// TIA Portal project "Delta_Praktika_P&P" (V17)

(* hardware
DEVICE "S7-1500/ET200MP station_1"  S7-1500 station
   slot 0: "Rail_0"  Rack  6ES7 590-1***0-0AA0
   slot 1: "PLC_2"  CPU 1517TF-3 PN/DP  6ES7 517-3UP00-0AB0  V2.9
      slot 3: "CPU display_1"  6ES7591-1BA00-0AA0
      slot 32768: "PROFINET interface_1"  X1
      slot 33024: "PROFINET interface_2"  X2
      slot 33280: "DP interface_1"  X3
      slot 34817: "Virtual CP interface port_1"  Virtual CP interface port  Virtual CP interface port
DEVICE "ET 200SP station_1"  ET 200SP-Station
   slot 0: "Rack_0"  Rack  6ES5 710-8MAx1
   slot 0: "et200sp"  IM 155-6 PN/2 HF  6ES7 155-6AU01-0CN0  V4.2
   slot 1: "DI 8x24VDC HF_1"  DI 8x24VDC HF  6ES7 131-6BF00-0CA0  V2.0
      slot 1: "DI 8x24VDC HF_1"  DI 8x24VDC HF
   slot 2: "DQ 8x24VDC/0.5A HF_1"  DQ 8x24VDC/0.5A HF  6ES7 132-6BF00-0CA0  V2.0
      slot 1: "DQ 8x24VDC/0.5A HF_1"  DQ 8x24VDC/0.5A HF
   slot 3: "CM 4xIO-Link_1"  CM 4xIO-Link  6ES7 137-6BD00-0BA0  V2.2
      slot 1: "CM 4xIO-Link_1"  6ES7 137-6BD00-0BA0
   slot 4: "Server module_1"  Server module  6ES7 193-6PA00-0AA0  V1.1
      slot 1: "Server module_1"  Server module
   slot 127: "BA 2xRJ45"  BA 2xRJ45  6ES7 193-6AR00-0AA0  V0.0
      slot 1: "Port_1"  X1 P1 R  6ES7 193-6AR00-0AA0  V0.0
      slot 2: "Port_2"  X1 P2 R  6ES7 193-6AR00-0AA0  V0.0
DEVICE "SINAMICS V_1"  SINAMICS V
   slot 0: "SINAMICS V90 PN Rack"  Rail  1.0
   slot 0: "a1"  V90 PN  6SL3 210-5FB10-4UFx  V1.4
      slot 1: "Drive object"  Drive Object
         slot 1: "Module access point"  Module Access Point
         slot 2: "Without PROFIsafe"  No ProfiSafe
         slot 3: "Telegram"  SIEMENS Telegramm 105
DEVICE "SINAMICS V_2"  SINAMICS V
   slot 0: "SINAMICS V90 PN Rack"  Rail  1.0
   slot 0: "a3"  V90 PN  6SL3 210-5FB10-4UFx  V1.4
      slot 1: "Drive object"  Drive Object
         slot 1: "Module access point"  Module Access Point
         slot 2: "Without PROFIsafe"  No ProfiSafe
         slot 3: "Telegram"  SIEMENS Telegramm 105
DEVICE "SINAMICS V_3"  SINAMICS V
   slot 0: "SINAMICS V90 PN Rack"  Rail  1.0
   slot 0: "a2"  V90 PN  6SL3 210-5FB10-4UFx  V1.4
      slot 1: "Drive object"  Drive Object
         slot 1: "Module access point"  Module Access Point
         slot 2: "Without PROFIsafe"  No ProfiSafe
         slot 3: "Telegram"  SIEMENS Telegramm 105
DEVICE "HMI_1"  KTP1200 Basic PN
   slot 0: "HMI_1"  KTP1200 Basic PN  6AV2 123-2MB03-0AX0  17.0.0.0
   slot 1: "HMI_RT_1"  KTP1200 Basic PN  6AV2 123-2MB03-0AX0  17.0.0.0
   slot 5: "HMI_1.IE_CP_1"  PROFINET Interface  17.0.0.0
      slot 1: "Interfaz PROFINET_1"  PROFINET Interface
         slot 1: "Port_1"  Port
*)

// ===== PLC "PLC_2"  CPU 1517TF-3 PN/DP =====

VAR_GLOBAL   // PLC tag table "Default tag table"
   "A1_Actor_Interface_AddressIn" AT %I0.0 : "PD_TEL3_IN";
   "A1_Actor_Interface_AddressOut" AT %Q0.0 : "PD_TEL3_OUT";
   "A2_Actor_Interface_AddressIn" AT %I18.0 : "PD_TEL3_IN";
   "A2_Actor_Interface_AddressOut" AT %Q10.0 : "PD_TEL3_OUT";
   "A3_Actor_Interface_AddressIn" AT %I36.0 : "PD_TEL3_IN";
   "A3_Actor_Interface_AddressOut" AT %Q20.0 : "PD_TEL3_OUT";
   "A1_axis_Actor_Interface_AddressIn" AT %I0.0 : "PD_TEL105_IN";
   "A1_axis_Actor_Interface_AddressOut" AT %Q0.0 : "PD_TEL105_OUT";
   "a2_axis_Actor_Interface_AddressIn" AT %I20.0 : "PD_TEL105_IN";
   "a2_axis_Actor_Interface_AddressOut" AT %Q63.0 : "PD_TEL105_OUT";
   "a3_asix_Actor_Interface_AddressIn" AT %I87.0 : "PD_TEL105_IN";
   "a3_asix_Actor_Interface_AddressOut" AT %Q83.0 : "PD_TEL105_OUT";
   "Freno_a1" AT %Q30.1 : Bool;
   "marka_Freno_a1" AT %M30.1 : Bool;
   "marka_Freno_a2" AT %M30.2 : Bool;
   "Freno_a2" AT %Q30.2 : Bool;
   "Freno_a3" AT %Q30.0 : Bool;
   "marka_Freno_a3" AT %M30.0 : Bool;
   "System_Byte" AT %MB256 : Byte;
   "FirstScan" AT %M256.0 : Bool;
   "DiagStatusUpdate" AT %M256.1 : Bool;
   "AlwaysTRUE" AT %M256.2 : Bool;
   "AlwaysFALSE" AT %M256.3 : Bool;
   "Clock_Byte" AT %MB255 : Byte;
   "Clock_10Hz" AT %M255.0 : Bool;
   "Clock_5Hz" AT %M255.1 : Bool;
   "Clock_2.5Hz" AT %M255.2 : Bool;
   "Clock_2Hz" AT %M255.3 : Bool;
   "Clock_1.25Hz" AT %M255.4 : Bool;
   "Clock_1Hz" AT %M255.5 : Bool;
   "Clock_0.625Hz" AT %M255.6 : Bool;
   "Clock_0.5Hz" AT %M255.7 : Bool;
   "Tag_1" AT %M401.0 : Bool;
   "JogFordward" AT %M150.0 : Bool;
   "JogBackward" AT %M150.1 : Bool;
   "Direction" AT %MB151 : USInt;
   "x+" AT %M152.0 : Bool;
   "x-" AT %M152.1 : Bool;
   "y+" AT %M152.2 : Bool;
   "y-" AT %M152.3 : Bool;
   "z+" AT %M152.4 : Bool;
   "z-" AT %M152.5 : Bool;
   "HABILITAR" AT %M150.2 : Bool;
   "Etapa0" AT %M0.0 : Bool;
   "HMI_start" AT %M10.0 : Bool;
   "Etapa1" AT %M0.1 : Bool;
   "Etapa2" AT %M0.2 : Bool;
   "Etapa3" AT %M0.3 : Bool;
   "Etapa4" AT %M0.4 : Bool;
   "Etapa5" AT %M0.5 : Bool;
   "Etapa6" AT %M0.6 : Bool;
   "Etapa7" AT %M0.7 : Bool;
   "kontagailua" AT %MW2 : Int;
   "Tag_2" AT %MB0 : Byte;
   "Tag_3" AT %M11.0 : Bool;
   "Etapa8" AT %M1.0 : Bool;
   "Etapa9" AT %M1.1 : Bool;
   "Etapa10" AT %M1.2 : Bool;
   "Etapa11" AT %M1.3 : Bool;
   "Etapa12" AT %M1.4 : Bool;
   "Tag_4" AT %MB1 : Byte;
   "Bentosa" AT %Q30.3 : Bool;
   "Tag_5" AT %M11.1 : Bool;
   "Tag_6" AT %M11.2 : Bool;
   "Tag_7" AT %M11.3 : Bool;
   "Tag_8" AT %M11.4 : Bool;
   "Tag_9" AT %M11.5 : Bool;
   "Tag_10" AT %M11.6 : Bool;
   "Tag_11" AT %M11.7 : Bool;
   "Tag_12" AT %M12.0 : Bool;
   "Tag_13" AT %M17.0 : Bool;
   "Tag_14" AT %M17.1 : Bool;
   "Tag_15" AT %M17.3 : Bool;
   "Tag_16" AT %M17.4 : Bool;
   "Tag_17" AT %M17.5 : Bool;
   "Tag_18" AT %M17.6 : Bool;
   "Tag_19" AT %M18.0 : Bool;
   "Tag_20" AT %M18.1 : Bool;
   "Tag_21" AT %M18.2 : Bool;
   "Tag_22" AT %M18.3 : Bool;
   "Tag_23" AT %M18.4 : Bool;
   "Tag_24" AT %M18.5 : Bool;
END_VAR

TYPE "LKinCtrl_typePathDynamics"
   STRUCT
      velocity : LReal := -1.0;   // >0.0: configured value used; <0.0: default TO setting used; for cmdType = 100 ==> waitTime in ms
      acceleration : LReal := -1.0;   // >0.0: configured value used; <0.0: default TO setting used
      deceleration : LReal := -1.0;   // >0.0: configured value used; <0.0: default TO setting used
      jerk : LReal := -1.0;   // >0.0: configured value used; <0.0: default TO setting used
   END_STRUCT;
END_TYPE

TYPE "LKinCtrl_typeSPTPDynamics"
   STRUCT
      velocityFactor : LReal;   // Factor for the velocity of axis movements in relation to the respective maximum velocity of the axes. Permitted value range: -1.0 < Factor ≤ 1.0
      accelerationFactor : LReal;   // Factor for the acceleration of axis movements in relation to the respective maximum acceleration of the axis. Permitted value range: -1.0 < Factor ≤ 1.0
      decelerationFactor : LReal;   // Factor for the deceleration of the axis movements in relation to the respective maximum deceleration of the axis. Permitted value range: -1.0 < Factor ≤ 1.0
      jerkFactor : LReal;   // Factor for the jerk of axis movements in relation to the respective maximum jerk of the axis. Permitted value range: -1.0 <Factor ≤ 0.0 and 0.1 < Factor ≤ 0.9
   END_STRUCT;
END_TYPE

TYPE "LKinCtrl_typeJogFrameDiagnostics"
VERSION : 0.1
// support: tech.team.motioncontrol@siemens.com
   STRUCT
      timeStamp : Date_And_Time;   // Time stamp at which the error occurred
      status : Word;   // Status of FB when error occurred
      stateNumber : DInt;   // State in the state machine of the FB when the error occurred
   END_STRUCT;
END_TYPE

TYPE "LKinCtrl_typeCartesianPosition"
   STRUCT
      x : LReal;   // X
      y : LReal;   // Y
      z : LReal;   // Z
      "a" : LReal;   // A
      "b" : LReal;   // B
      c : LReal;   // C
   END_STRUCT;
END_TYPE

TYPE "LKinCtrl_typeDynamics"
VERSION : 0.1
   STRUCT
      path : "LKinCtrl_typePathDynamics";   // Specification of the path dynamics
      orientation : "LKinCtrl_typePathDynamics";   // Specification of the orientation dynamics
      dynamicAdaption : DInt := 1;   // 0=no dynamic adaption, 1=dynamic adaptation with segmentation of the path, 2=dynamic adaptation without segmentation of the path
      directionA : DInt := 3;   // 1=positive direction, 2=negative direction, 3=shortest distance
      sPTP : "LKinCtrl_typeSPTPDynamics";   // Specification of the dynamic factor for sptp movement
   END_STRUCT;
END_TYPE

DATA_BLOCK "Power_DB"   // DB9
{ S7_Optimized_Access := 'TRUE' }
VERSION : 0.1
// stored: InstanceOfName Power
"Power"
BEGIN
END_DATA_BLOCK

DATA_BLOCK "Parametroak"   // DB11
{ S7_Optimized_Access := 'TRUE' }
VERSION : 0.1
   VAR
      Abiadura : LReal := 2.0;
      Azelerazioa : LReal := 40.0;
      Desazelerazioa : LReal := 40.0;
      Jerk : LReal := 400.0;
      offset : LReal := 30.0;
   END_VAR
BEGIN
END_DATA_BLOCK

DATA_BLOCK "Jog_DB"   // DB14
{ S7_Optimized_Access := 'TRUE' }
VERSION : 0.1
// stored: InstanceOfName Jog
"Jog"
BEGIN
END_DATA_BLOCK

DATA_BLOCK "Hominga_DB"   // DB18
{ S7_Optimized_Access := 'TRUE' }
VERSION : 0.1
// stored: InstanceOfName Hominga
"Hominga"
BEGIN
END_DATA_BLOCK

DATA_BLOCK "Puntuak"   // DB24
{ S7_Optimized_Access := 'TRUE' }
VERSION : 0.1
   VAR
      Puntu_abs_home : Array[1..4] of LReal;
      Puntu_abs_1 : Array[1..4] of LReal;
      Puntu_abs_2 : Array[1..4] of LReal;
      Puntu_rel_1 : Array[1..4] of LReal;
      Puntu_aux_1 : Array[1..3] of LReal;
      Puntu_zirkular_1 : Array[1..4] of LReal;
      HMI_erlatibo_lineal : Array[1..4] of LReal;
      HMI_abs_lineal : Array[1..4] of LReal;
      HMI_abs_zirkular_aux : Array[1..3] of LReal;
      HMI_abs_zirkular_endpoint : Array[1..4] of LReal;
      HMI_abs_ptp : Array[1..4] of LReal;
   END_VAR
BEGIN
   Puntu_abs_home[1] := 0.0;
   Puntu_abs_home[2] := 0.0;
   Puntu_abs_home[3] := -722.59;
   Puntu_abs_home[4] := 0.0;
   Puntu_abs_1[1] := 0.0;
   Puntu_abs_1[2] := 0.0;
   Puntu_abs_1[3] := -700.0;
   Puntu_abs_1[4] := 0.0;
   Puntu_rel_1[1] := 50.0;
   Puntu_rel_1[2] := 0.0;
   Puntu_rel_1[3] := 0.0;
   Puntu_abs_2[1] := 50.0;
   Puntu_abs_2[2] := 50.0;
   Puntu_abs_2[3] := -700.0;
   Puntu_abs_2[4] := 0.0;
   Puntu_aux_1[1] := 50.0;
   Puntu_aux_1[2] := 0.0;
   Puntu_aux_1[3] := -700.0;
   Puntu_zirkular_1[1] := 100.0;
   Puntu_zirkular_1[2] := 0.0;
   Puntu_zirkular_1[3] := -700.0;
   Puntu_zirkular_1[4] := 0.0;
END_DATA_BLOCK

DATA_BLOCK "ParametroakII"   // DB25
{ S7_Optimized_Access := 'TRUE' }
VERSION : 0.1
   VAR
      abiadura : LReal := 10.0;
      azelerazioa : LReal := 20.0;
      desazelerazioa : LReal := 20.0;
      jerk : LReal := 40.0;
   END_VAR
BEGIN
END_DATA_BLOCK

DATA_BLOCK "LKinCtrl_MC_JogFrame_DB"   // DB30
{ S7_Optimized_Access := 'TRUE' }
AUTHOR : tech.team.motioncontrol@siemens.com
FAMILY : LKinCtrl
VERSION : 1.1
// stored: InstanceOfName LKinCtrl_MC_JogFrame
"LKinCtrl_MC_JogFrame"
BEGIN
END_DATA_BLOCK

DATA_BLOCK "LKinCtrl_MC_JogFrame_DB_1"   // DB31
{ S7_Optimized_Access := 'TRUE' }
AUTHOR : tech.team.motioncontrol@siemens.com
FAMILY : LKinCtrl
VERSION : 1.1
// stored: InstanceOfName LKinCtrl_MC_JogFrame
"LKinCtrl_MC_JogFrame"
BEGIN
END_DATA_BLOCK

DATA_BLOCK "Delta_robota_ajusteak"   // DB32
{ S7_Optimized_Access := 'TRUE' }
VERSION : 0.1
   VAR
      Jog_aldagaiak : "LKinCtrl_typeDynamics";
   END_VAR
BEGIN
   Jog_aldagaiak.path.velocity := 10.0;
   Jog_aldagaiak.path.acceleration := 20.0;
   Jog_aldagaiak.path.deceleration := 20.0;
   Jog_aldagaiak.path.jerk := 40.0;
END_DATA_BLOCK

DATA_BLOCK "PickandPlace"   // DB33
{ S7_Optimized_Access := 'TRUE' }
VERSION : 0.1
   VAR
      P11 : Array[1..4] of LReal;
      P12 : Array[1..4] of LReal;
      P13 : Array[1..4] of LReal;
      P14 : Array[1..4] of LReal;
      P15 : Array[1..4] of LReal;
      P16 : Array[1..4] of LReal;
      P21 : Array[1..4] of LReal;
      P22 : Array[1..4] of LReal;
      P23 : Array[1..4] of LReal;
      P24 : Array[1..4] of LReal;
      P25 : Array[1..4] of LReal;
      P26 : Array[1..4] of LReal;
      HOME_Maketa : Array[1..4] of LReal;
      HOME_Prozesua : Array[1..4] of LReal;
      "Puntu_PiezaZ+" : Array[1..4] of LReal;
      Puntu_Pieza : Array[1..4] of LReal;
   END_VAR
BEGIN
   P11[1] := -4.015;
   P11[2] := 149.099;
   P11[3] := -636.999;
   P12[1] := -40.434;
   P12[2] := 134.412;
   P12[3] := -638.334;
   P13[1] := -1.376;
   P13[2] := 111.506;
   P13[3] := -651.752;
   P14[1] := -37.504;
   P14[2] := 99.396;
   P14[3] := -651.9;
   P15[1] := 0.409;
   P15[2] := 70.62;
   P15[3] := -662.979;
   P16[1] := -35.408;
   P16[2] := 60.504;
   P16[3] := -663.138;
   P21[1] := 32.325;
   P21[2] := -88.2;
   P21[3] := -658.347;
   P22[1] := -1.0;
   P22[2] := -89.9;
   P22[3] := -658.633;
   P23[1] := 42.333;
   P23[2] := -127.0;
   P23[3] := -644.987;
   P24[1] := 8.91;
   P24[2] := -127.925;
   P24[3] := -645.448;
   P25[1] := 52.87;
   P25[2] := -166.925;
   P25[3] := -625.259;
   P26[1] := 21.0;
   P26[2] := -166.0;
   P26[3] := -627.242;
   HOME_Maketa[1] := 0.0;
   HOME_Maketa[2] := 0.0;
   HOME_Maketa[3] := -722.59;
   HOME_Maketa[4] := 0.0;
   HOME_Prozesua[1] := 0.0;
   HOME_Prozesua[2] := 0.0;
   HOME_Prozesua[3] := -700.0;
   HOME_Prozesua[4] := 0.0;
END_DATA_BLOCK

// folder: System blocks/Program resources

DATA_BLOCK "IEC_Timer_0_DB"   // DB36
{ S7_Optimized_Access := 'TRUE' }
AUTHOR : Simatic
FAMILY : IEC
NAME : IEC_TMR
VERSION : 1.0
// stored: InstanceOfName IEC_TIMER
"IEC_TIMER"
BEGIN
END_DATA_BLOCK

DATA_BLOCK "IEC_Timer_0_DB_1"   // DB37
{ S7_Optimized_Access := 'TRUE' }
AUTHOR : Simatic
FAMILY : IEC
NAME : IEC_TMR
VERSION : 1.0
// stored: InstanceOfName IEC_TIMER
"IEC_TIMER"
BEGIN
END_DATA_BLOCK

DATA_BLOCK "IEC_Timer_0_DB_2"   // DB39
{ S7_Optimized_Access := 'TRUE' }
AUTHOR : Simatic
FAMILY : IEC
NAME : IEC_TMR
VERSION : 1.0
// stored: InstanceOfName IEC_TIMER
"IEC_TIMER"
BEGIN
END_DATA_BLOCK

DATA_BLOCK "IEC_Timer_0_DB_3"   // DB40
{ S7_Optimized_Access := 'TRUE' }
AUTHOR : Simatic
FAMILY : IEC
NAME : IEC_TMR
VERSION : 1.0
// stored: InstanceOfName IEC_TIMER
"IEC_TIMER"
BEGIN
END_DATA_BLOCK

DATA_BLOCK "IEC_Timer_0_DB_4"   // DB41
{ S7_Optimized_Access := 'TRUE' }
AUTHOR : Simatic
FAMILY : IEC
NAME : IEC_TMR
VERSION : 1.0
// stored: InstanceOfName IEC_TIMER
"IEC_TIMER"
BEGIN
END_DATA_BLOCK

// folder: (top level)

DATA_BLOCK "a1_asix"   // DB2, Motion_DB
{ S7_Optimized_Access := 'TRUE' }
AUTHOR : SIMATIC
FAMILY : MC_1500
VERSION : 6.0
// stored: InstanceOfName TO_PositioningAxis
"TO_PositioningAxis"
BEGIN
END_DATA_BLOCK

DATA_BLOCK "a2_axis"   // DB3, Motion_DB
{ S7_Optimized_Access := 'TRUE' }
AUTHOR : SIMATIC
FAMILY : MC_1500
VERSION : 6.0
// stored: InstanceOfName TO_PositioningAxis
"TO_PositioningAxis"
BEGIN
END_DATA_BLOCK

DATA_BLOCK "a3_axis"   // DB4, Motion_DB
{ S7_Optimized_Access := 'TRUE' }
AUTHOR : SIMATIC
FAMILY : MC_1500
VERSION : 6.0
// stored: InstanceOfName TO_PositioningAxis
"TO_PositioningAxis"
BEGIN
END_DATA_BLOCK

DATA_BLOCK "Delta_Robota"   // DB7, Motion_DB
{ S7_Optimized_Access := 'TRUE' }
AUTHOR : SIMATIC
FAMILY : MC_1500
VERSION : 6.0
// stored: InstanceOfName TO_Kinematics
"TO_Kinematics"
BEGIN
END_DATA_BLOCK

FUNCTION_BLOCK "Power"   // FB2, LAD
{ S7_Optimized_Access := 'TRUE' }
VERSION : 0.1
   VAR_INPUT
      Power_a1 : Bool;
      Power_a2 : Bool;
      Power_a3 : Bool;
   END_VAR
   VAR_OUTPUT
      Status_a1 : Bool;
      Status_a2 : Bool;
      Status_a3 : Bool;
      Error_a1 : Bool;
      Error_a2 : Bool;
      Error_a3 : Bool;
   END_VAR
BEGIN

REGION Network 1
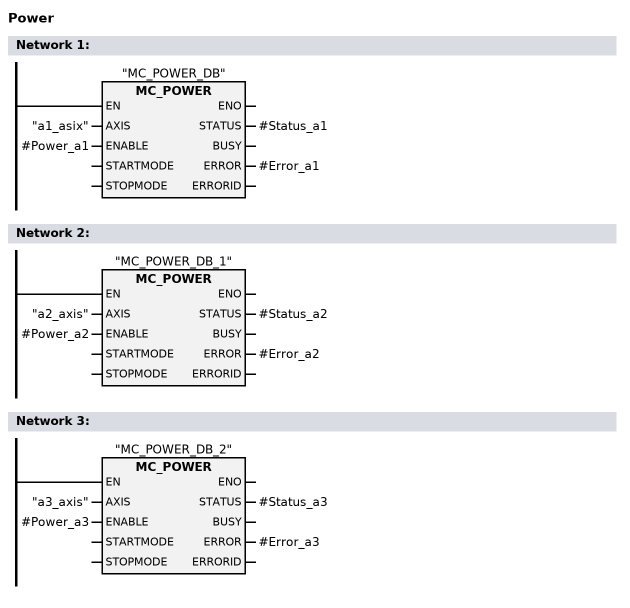
   "MC_POWER_DB"(Axis := "a1_asix", Enable := #Power_a1, Status => #Status_a1, Error => #Error_a1);   // MC_POWER
END_REGION

REGION Network 2
   "MC_POWER_DB_1"(Axis := "a2_axis", Enable := #Power_a2, Status => #Status_a2, Error => #Error_a2);   // MC_POWER
END_REGION

REGION Network 3
   "MC_POWER_DB_2"(Axis := "a3_axis", Enable := #Power_a3, Status => #Status_a3, Error => #Error_a3);   // MC_POWER
END_REGION
END_FUNCTION_BLOCK

FUNCTION_BLOCK "Jog"   // FB3, LAD
{ S7_Optimized_Access := 'TRUE' }
VERSION : 0.1
   VAR_INPUT
      "A1+" : Bool;
      "A1-" : Bool;
      "A2+" : Bool;
      "A2-" : Bool;
      "A3+" : Bool;
      "A3-" : Bool;
   END_VAR
BEGIN

REGION Network 1
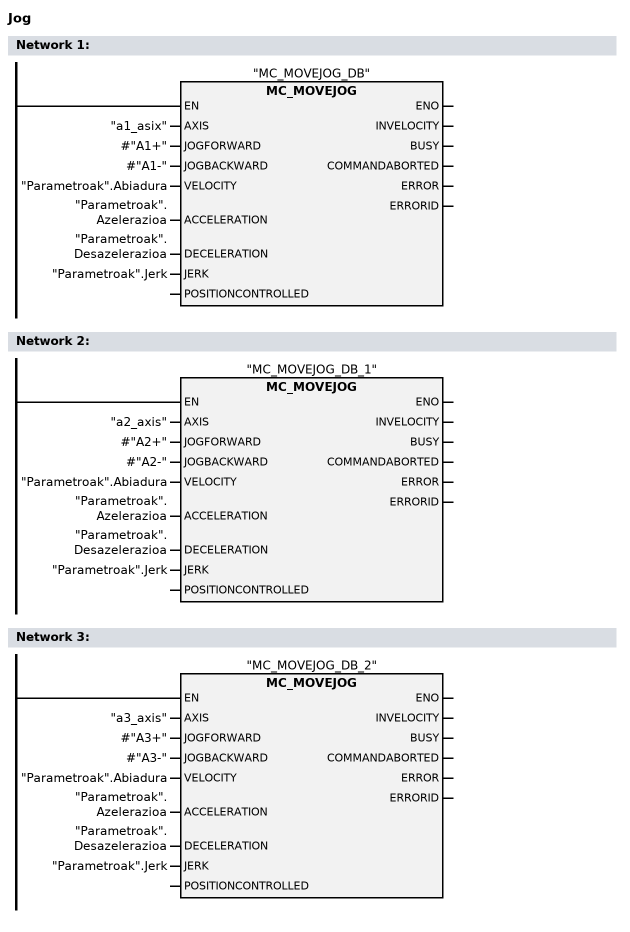
   "MC_MOVEJOG_DB"(Axis := "a1_asix",   // MC_MOVEJOG
                   JogForward := #"A1+",
                   JogBackward := #"A1-",
                   Velocity := "Parametroak".Abiadura,
                   Acceleration := "Parametroak".Azelerazioa,
                   Deceleration := "Parametroak".Desazelerazioa,
                   Jerk := "Parametroak".Jerk);
END_REGION

REGION Network 2
   "MC_MOVEJOG_DB_1"(Axis := "a2_axis",   // MC_MOVEJOG
                     JogForward := #"A2+",
                     JogBackward := #"A2-",
                     Velocity := "Parametroak".Abiadura,
                     Acceleration := "Parametroak".Azelerazioa,
                     Deceleration := "Parametroak".Desazelerazioa,
                     Jerk := "Parametroak".Jerk);
END_REGION

REGION Network 3
   "MC_MOVEJOG_DB_2"(Axis := "a3_axis",   // MC_MOVEJOG
                     JogForward := #"A3+",
                     JogBackward := #"A3-",
                     Velocity := "Parametroak".Abiadura,
                     Acceleration := "Parametroak".Azelerazioa,
                     Deceleration := "Parametroak".Desazelerazioa,
                     Jerk := "Parametroak".Jerk);
END_REGION
END_FUNCTION_BLOCK

FUNCTION_BLOCK "Hominga"   // FB4, LAD
{ S7_Optimized_Access := 'TRUE' }
VERSION : 0.1
   VAR_INPUT
      homing_a1 : Bool;
      homing_a2 : Bool;
      homing_a3 : Bool;
   END_VAR
   VAR_OUTPUT
      Done_a1 : Bool;
      Done_a2 : Bool;
      Done_a3 : Bool;
   END_VAR
BEGIN

REGION Network 1
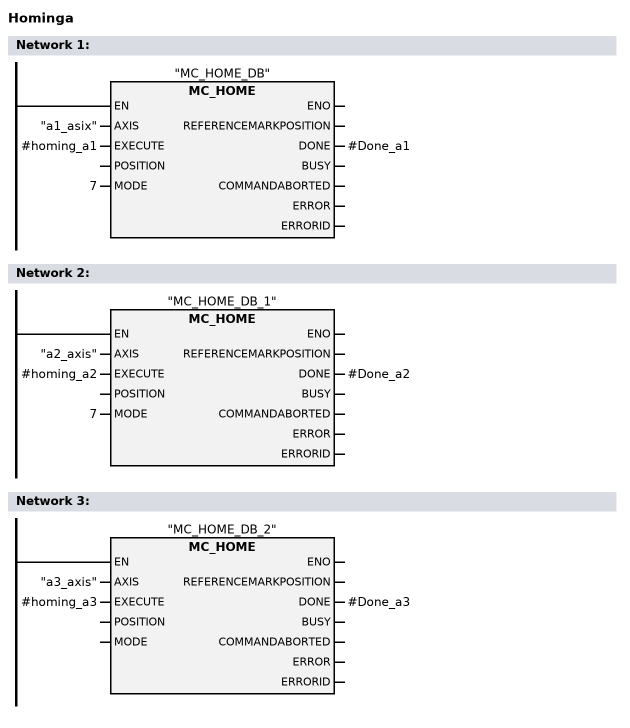
   "MC_HOME_DB"(Axis := "a1_asix", Execute := #homing_a1, Mode := 7, Done => #Done_a1);   // MC_HOME
END_REGION

REGION Network 2
   "MC_HOME_DB_1"(Axis := "a2_axis", Execute := #homing_a2, Mode := 7, Done => #Done_a2);   // MC_HOME
END_REGION

REGION Network 3
   "MC_HOME_DB_2"(Axis := "a3_axis", Execute := #homing_a3, Done => #Done_a3);   // MC_HOME
END_REGION
END_FUNCTION_BLOCK

FUNCTION_BLOCK "LKinCtrl_MC_JogFrame"   // FB35010, SCL
TITLE = LKinCtrl_MC_JogFrame
{ S7_Optimized_Access := 'TRUE' }
AUTHOR : tech.team.motioncontrol@siemens.com
FAMILY : LKinCtrl
VERSION : 1.1
// Functionality: This function block provides various jog functionality for kinematics technology object.
   VAR_INPUT
      jogForward : Bool := FALSE;   // Jog the kinematics forward in the selected jog direction
      jogBackward : Bool := FALSE;   // Jog the kinematics backward in the selected jog direction
      jogToPosition : Bool := FALSE;   // Jog the kinematics to the specified target position
      jogSPTP : Bool := FALSE;   // Jog the kinematics synchronous point to point
      jogDirection : USInt := 1;   // 1=x-direction, 2=y-direction, 3=z-direction, 4=a-direction
      jogModeInc : Bool := FALSE;   // 1=incremental jog mode, 0=continuous jog mode
      jogIncrement : LReal := 1.0;   // Specification of the jog increment
      targetPosition : "LKinCtrl_typeCartesianPosition";   // Specification of the target position
      coordSystem : DInt := 0;   // 0=WCS, 1= OCS1, 2=OCS2, 3=OCS3, 100=MCS
      linkconstellation : DWord := 16#FFFF_FFFF;   // Target joint position space
      tool : DInt := 1;   // 1= tool1, 2=tool2, 3=tool3
      dynamics : "LKinCtrl_typeDynamics";   // Specification of the jog dynamics
   END_VAR
   VAR_OUTPUT
      done : Bool := FALSE;   // TRUE: Commanded functionality has been completed successfully
      busy : Bool := FALSE;   // TRUE: FB is not finished and new output values can be expected
      active : Bool := FALSE;   // TRUE: The setpoints are calculated
      error : Bool := FALSE;   // TRUE: An error occurred during the execution of the FB
      status : Word := 16#7000;   // 16#0000 - 16#7FFF: Status of the FB, 16#8000 - 16#FFFF: Error identification
      remainingDistance : LReal := 0.0;   // Distance-to-go of the current job
      diagnostics : "LKinCtrl_typeJogFrameDiagnostics";   // Diagnostics information
   END_VAR
   VAR_IN_OUT
      axesGroup : TO_Kinematics;   // Kinematics technology object
   END_VAR
   VAR
      instMC_SetTool : MC_SETTOOL;   // Instance MC_SetTool
      instMC_GroupStop : MC_GROUPSTOP;   // Instance MC_GroupStop
      instMC_MoveLinearAbsoute : MC_MOVELINEARABSOLUTE;   // Instance MC_MoveLinearAbsolute
      instMC_MoveLinearRelative : MC_MOVELINEARRELATIVE;   // Instance MC_MoveLinearRelative
      instMC_MoveDirectAbsolute : MC_MOVEDIRECTABSOLUTE;   // Instance MC_MoveDirectAbsolute
      statDone : Bool := FALSE;   // Static value for output 'done'
      statBusy : Bool := FALSE;   // Static value for output 'busy'
      statActive : Bool := FALSE;   // Static value for output 'active'
      statError : Bool := FALSE;   // Static value for output 'error'
      statStatus : Word := 16#7000;   // 0000=STATUS_EXECUTION_FINISHED; 7000=STATUS_NO_CALL; 7001=STATUS_FIRST_CALL; 7002=STATUS_SUBSEQUENT_CALL; 8600=ERR_UNDEFINED_STATE
      statRemainingDistance : LReal := 0.0;   // Static value for remaining distance
      statFBState : DInt := 0;   // 0= NO PROCESSING; 10=IDLE; 20=SET_TOOL; 30=SET_DYNAMICS, 50=EXECUTE_MOVEMENT; 100=STOP
      statToolOld : DInt := 1;   // Static value for tool
      statJogForwardOld : Bool := FALSE;   // Static value for jog forward command
      statJogBackwardOld : Bool := FALSE;   // Static value for jog backward command
      statJogToPositionOld : Bool := FALSE;   // Static value for jog to position command
      statJogSPTPOld : Bool := FALSE;   // Static value for jog sPTP command
      statOrientationDynamicsChanged : Bool := FALSE;   // Static value indicates that default orientation dynamics have been changed
      statOrientationDynamicsOld : "LKinCtrl_typePathDynamics";   // Static value for orientation dynamics
   END_VAR
   VAR_TEMP
      tempJogForward : Bool;   // Temporary variable for jog forward input
      tempJogBackward : Bool;   // Temporary variable for jog backward input
      tempJogToPosition : Bool;   // Temporary variable for jog to position input
      tempJogSPTP : Bool;   // Temporary variable for jog sptp input
      tempCounter : DInt;   // Temporary variable for counter
      tempRet : Int;   // Temporary variable for time stamp if error occurred
   END_VAR
   VAR CONSTANT
      FB_STATE_NO_PROCESSING : DInt := 0;   // FB state: No processing
      FB_STATE_CMD_CONFIGURATION : DInt := 10;   // FB state: Basic command configuration are set depending on input parameter
      FB_STATE_SET_TOOL : DInt := 20;   // FB state: Tool change is performed if required
      FB_STATE_EXECUTE_MOVEMENT : DInt := 50;   // FB state: Command is being executed
      FB_STATE_STOP : DInt := 100;   // FB state: Kinematics movement is stopped
      STATUS_EXECUTION_FINISHED : Word := 16#0000;   // The command execution is finished by reaching the target position or stopping the jog command
      STATUS_NO_CALL : Word := 16#7000;   // No call of FB
      STATUS_FIRST_CALL : Word := 16#7001;   // First cycle of FB after enabling
      STATUS_SUBSEQUENT_CALL : Word := 16#7002;   // FB enabled
      ERR_UNDEFINED_STATE : Word := 16#8600;   // Error due to an undefined FB state
      ERR_TO_KINEMATICS : Word := 16#8001;   // Error at technology object kinematics
      ERR_INVALID_JOG_DIRECTION : Word := 16#8007;   // The specified jog direction is invalid (valid values are 1=x-direction, 2=y-direction, 3=z-direction, 4=a-direction)
      ERR_MOTION_JOB_IN_PROGRESS : Word := 16#8090;   // A motion job is in progress or the kinematics control panel is activated
      ERR_TWO_JOG_COMMANDS_SIMULTANEOUSLY : Word := 16#8091;   // Two jog commands were triggered simultaneously
      ERR_INVALID_COORDINATE_SYSTEM : Word := 16#80B1;   // The specified coordinate system is invalid (valid values are 0=WCS, 1= OCS1, 2=OCS2, 3=OCS3)
      ERR_INVALID_TOOL : Word := 16#80CA;   // The specified tool is invalid (valid values are 1= tool1, 2=tool2, 3=tool3)
      MAX_DISTANCE : LReal := 700000000.0;   // The value is set for relative linear movement as jog increment for icremental jog mode
      L_BOUND_TOOL : DInt := 1;   // Lower bound for tool selection
      U_BOUND_TOOL : DInt := 3;   // Upper bound for tool selection
      L_BOUND_JOG_DIRECTION : DInt := 1;   // Lower bound for jog direction selection
      U_BOUND_JOG_DIRECTION : DInt := 4;   // Upper bound for jog direction selection
      L_BOUND_COORDSYSTEM : DInt := 0;   // Lower bound for coordinate system selection
      U_BOUND_COORDSYSTEM : DInt := 3;   // Upper bound for coordinate system selection
      INDEX_COORDSYSTEM_MCS : DInt := 100;   // Coordinate system index for MCS
   END_VAR
   // dynamics.sPTP.velocityFactor := -1.0;
   // dynamics.sPTP.accelerationFactor := -1.0;
   // dynamics.sPTP.decelerationFactor := -1.0;
   // dynamics.sPTP.jerkFactor := -1.0;
BEGIN
   //=============================================================================
   // SIEMENS AG
   // (c)Copyright 2018 All Rights Reserved
   //-----------------------------------------------------------------------------
   // Library:       LKinCtrl
   // Tested with:   S7-1516T
   // Engineering:   TIA Portal V15
   // Restrictions:  -
   // Requirements:  S7-1500T FW 2.5
   // Functionality: LKinCtrl_MC_JogFrame
   // This function block provides various jog functionality for kinematics technology object
   // 
   // Support: tech.team.motioncontrol@siemens.com
   // Note: Parameter comments are only available in language 'English (United States)'
   //-----------------------------------------------------------------------------
   // Change log table:
   // Version  Date        Expert in charge   Changes applied
   // 01.00.00 05.04.2018  IP                 First released version
   // 01.00.01 24.04.2018  IP                 Hotfix - initialization - no functional changes
   // 01.01.00 31.07.2018  IP                 Adjustment of input validation
   //                                         New wait condition for next movement until stopping is done
   //                                         Additional output parameter active and remaining distance
   // 01.01.01 07.08.2018  IP                 Hotfix - constant MAX_DISTANCE decreased
   // 01.01.02 09.01.2019  IP                 Hotfix - error indification adjusted
   // 01.01.03 14.01.2019  IP                 Hotfix - dynamics configuration adjusted
   // 01.01.04 12.07.2021  FF                 Added Synchronous point to point jogging
   // 01.01.05 14.12.2021  FR                 Fix for orientation dynamics and refactor
   // 01.01.06 15.07.2022  FR                 Fix for Override = 0 and fast toggle of inputs
   //=============================================================================

   #tempJogForward := #jogForward; // Work with temporary value / create process image
   #tempJogBackward := #jogBackward;
   #tempJogToPosition := #jogToPosition;
   #tempJogSPTP := #jogSPTP;

   REGION TRIGGERING

     IF ((#tempJogForward AND NOT #statJogForwardOld) // Check if FB is triggered
       OR (#tempJogBackward AND NOT #statJogBackwardOld)
       OR (#tempJogToPosition AND NOT #statJogToPositionOld)
       OR (#tempJogSPTP AND NOT #statJogSPTPOld))
       AND (#statStatus = #STATUS_NO_CALL)
       AND (#statFBState = #FB_STATE_NO_PROCESSING)
     THEN

       // First call; set FB variables for outputs
       #statBusy := TRUE;
       #statDone := FALSE;
       #statActive := FALSE;
       #statError := FALSE;
       #statRemainingDistance := 0.0;
       #statStatus := #STATUS_FIRST_CALL;

       // check if input parameter are valid
       IF (#jogDirection < #L_BOUND_JOG_DIRECTION OR #jogDirection > #U_BOUND_JOG_DIRECTION) // check jog direction
         AND (NOT #tempJogToPosition OR NOT #tempJogSPTP) THEN
         #statStatus := #ERR_INVALID_JOG_DIRECTION;
       ELSIF #tool < #L_BOUND_TOOL OR #tool > #U_BOUND_TOOL THEN // check tool
         #statStatus := #ERR_INVALID_TOOL;
       ELSIF (#coordSystem < #L_BOUND_COORDSYSTEM OR #coordSystem > #U_BOUND_COORDSYSTEM)
         AND NOT (#tempJogSPTP AND #coordSystem = #INDEX_COORDSYSTEM_MCS) // Double check for sPTP
       THEN // check coordinate system
         #statStatus := #ERR_INVALID_COORDINATE_SYSTEM;
       ELSIF NOT #axesGroup.StatusWord.%X6 THEN // check if a motion job is in progress or the kinematics control panel is activated
         #statStatus := #ERR_MOTION_JOB_IN_PROGRESS;
       ELSE // all input parameter are valid

         // reset execute inputs
         #instMC_GroupStop.Execute := FALSE;
         #instMC_MoveLinearAbsoute.Execute := FALSE;
         #instMC_MoveLinearRelative.Execute := FALSE;
         #instMC_MoveDirectAbsolute.Execute := FALSE;
         #instMC_SetTool.Execute := FALSE;

         // call FBs with execute = false
         #instMC_GroupStop(AxesGroup := #axesGroup);
         #instMC_MoveLinearAbsoute(AxesGroup := #axesGroup);
         #instMC_MoveLinearRelative(AxesGroup := #axesGroup);
         #instMC_MoveDirectAbsolute(AxesGroup := #axesGroup);
         #instMC_SetTool(AxesGroup := #axesGroup);

         // get actual tool number
         #statToolOld := #axesGroup.StatusTool.ActiveTool;

         // safe default dynamics for orientation axis
         #statOrientationDynamicsOld.velocity := #axesGroup.DynamicDefaults.Orientation.Velocity;
         #statOrientationDynamicsOld.acceleration := #axesGroup.DynamicDefaults.Orientation.Acceleration;
         #statOrientationDynamicsOld.deceleration := #axesGroup.DynamicDefaults.Orientation.Deceleration;
         #statOrientationDynamicsOld.jerk := #axesGroup.DynamicDefaults.Orientation.Jerk;
         #statOrientationDynamicsChanged := FALSE;

         // state machine - start functionality
         #statFBState := #FB_STATE_CMD_CONFIGURATION;
       END_IF;

     ELSIF (#statStatus = #STATUS_FIRST_CALL) THEN
       #statStatus := #STATUS_SUBSEQUENT_CALL;
     END_IF;

   END_REGION TRIGGERING

   IF (#statStatus = #STATUS_NO_CALL) THEN // Nothing to do -> End here to reduce "system load"
     RETURN;
   END_IF;

   REGION STOP_MOTION
     // detection of falling edge on jog command
     IF ((NOT #tempJogForward AND #statJogForwardOld)
       OR (NOT #tempJogBackward AND #statJogBackwardOld)
       OR (NOT #tempJogToPosition AND #statJogToPositionOld)
       OR (NOT #tempJogSPTP AND #statJogSPTPOld))
       AND NOT (#statFBState = #FB_STATE_NO_PROCESSING)
     THEN // stop jog command
       #statFBState := #FB_STATE_STOP;

       // two jog commands simultaneously    
     ELSIF ((#tempJogBackward AND #tempJogForward)
       OR (#tempJogBackward AND #tempJogToPosition)
       OR (#tempJogBackward AND #tempJogSPTP)
       OR (#tempJogForward AND #tempJogToPosition)
       OR (#tempJogForward AND #tempJogSPTP)
       OR (#tempJogToPosition AND #tempJogSPTP))
       AND NOT (#statFBState = #FB_STATE_NO_PROCESSING)
     THEN // stop jog command
       #statFBState := #FB_STATE_STOP;
       #statStatus := #ERR_TWO_JOG_COMMANDS_SIMULTANEOUSLY;
     END_IF;

     IF #statStatus <> #STATUS_FIRST_CALL AND (#statStatus.%X15 = FALSE) THEN
       IF #axesGroup.StatusWord.%X1 // general TO error
         OR #instMC_MoveLinearRelative.Error
         OR #instMC_GroupStop.Error
         OR #instMC_MoveLinearAbsoute.Error
         OR #instMC_MoveDirectAbsolute.Error
         OR #instMC_SetTool.Error
       THEN
         #statFBState := #FB_STATE_STOP;
       END_IF;
     END_IF;

   END_REGION

   // Edge detection 'execute' input
   #statJogForwardOld := #tempJogForward;
   #statJogBackwardOld := #tempJogBackward;
   #statJogToPositionOld := #tempJogToPosition;
   #statJogSPTPOld := #tempJogSPTP;

   REGION RESET_DEFAULT_ORIENTATION_DYNAMICS

     IF (#instMC_MoveLinearRelative.Busy OR #instMC_MoveLinearAbsoute.Busy OR #statFBState = #FB_STATE_STOP)
       AND #statOrientationDynamicsChanged
     THEN // reset default orientation dynamics
       #axesGroup.DynamicDefaults.Orientation.Velocity := #statOrientationDynamicsOld.velocity;
       #axesGroup.DynamicDefaults.Orientation.Acceleration := #statOrientationDynamicsOld.acceleration;
       #axesGroup.DynamicDefaults.Orientation.Deceleration := #statOrientationDynamicsOld.deceleration;
       #axesGroup.DynamicDefaults.Orientation.Jerk := #statOrientationDynamicsOld.jerk;
       #statOrientationDynamicsChanged := FALSE;
     END_IF;

   END_REGION

   REGION ACTIVE_OUTPUT

     // set active output if any of motion commands is active
     #statActive := #instMC_MoveLinearAbsoute.Active OR #instMC_MoveLinearRelative.Active OR #instMC_MoveDirectAbsolute.Active OR #instMC_GroupStop.Active;

   END_REGION

   REGION REMAINING_DISTANCE

     // set remaining distance at output if incremental mode active or while jogging to target position
     IF #instMC_MoveLinearAbsoute.Busy THEN
       #statRemainingDistance := #instMC_MoveLinearAbsoute.RemainingDistance;
     ELSIF #instMC_MoveLinearRelative.Busy AND #jogModeInc THEN
       #statRemainingDistance := #instMC_MoveLinearRelative.RemainingDistance;
     ELSE
       #statRemainingDistance := 0.0;
     END_IF;

   END_REGION

   REGION STATE_MACHINE

     CASE #statFBState OF // State machine of FB
       #FB_STATE_NO_PROCESSING: // No processing active (Note: this state must always be present and left empty)
         ;

       #FB_STATE_CMD_CONFIGURATION:
         // Check for override <> 0 -> Only execute commands if override <> 0 as there are issues with TO_Kin if override = 0
         IF #axesGroup.Override.Velocity <> 0 THEN

           REGION CONFIGURATION

             // jog forward or backward
             //*********************************************************************************************************
             IF #tempJogForward OR #tempJogBackward THEN
               // set MC_MoveLinearRelative parameter
               #instMC_MoveLinearRelative.CoordSystem := #coordSystem;
               #instMC_MoveLinearRelative.Velocity := #dynamics.path.velocity;
               #instMC_MoveLinearRelative.Acceleration := #dynamics.path.acceleration;
               #instMC_MoveLinearRelative.Deceleration := #dynamics.path.deceleration;
               #instMC_MoveLinearRelative.Jerk := #dynamics.path.jerk;

               // initialize jog distance - clear old values
               FOR #tempCounter := 1 TO 4 DO
                 #instMC_MoveLinearRelative.Distance[#tempCounter] := 0.0;
               END_FOR;

               // set jog mode
               IF #jogModeInc THEN // incremental
                 IF #tempJogForward THEN
                   #instMC_MoveLinearRelative.Distance[#jogDirection] := #jogIncrement;
                 ELSIF #tempJogBackward THEN
                   #instMC_MoveLinearRelative.Distance[#jogDirection] := - #jogIncrement;
                 END_IF;
                 #instMC_MoveLinearRelative.DynamicAdaption := #dynamics.dynamicAdaption;

               ELSE // continouos
                 IF #tempJogForward THEN
                   #instMC_MoveLinearRelative.Distance[#jogDirection] := #MAX_DISTANCE;
                 ELSIF #tempJogBackward THEN
                   #instMC_MoveLinearRelative.Distance[#jogDirection] := - #MAX_DISTANCE;
                 END_IF;

                 // switch off dynamic adaption for continouos mode
                 #instMC_MoveLinearRelative.DynamicAdaption := 0;
               END_IF;